VERSION : 1.1
// The function calculates a contour offset of a path (tool length and radius) / The function calculates a contour offset of a path (tool length and radius offset)
   VAR_INPUT
      toolLength : LReal;   // Tool length
      toolRadius : LReal;   // Tool radius
      pathPlane : Int;   // Path plane: XZ= 0, YZ=1, XY= 2
      compensationDirection : Int;   // Tool radius compensation direction: left=1, right = 0
   END_VAR
   VAR_IN_OUT
      pathDataIn : "LKinCtrl_typeCOffPathDataIn";   // Path data in
      pathDataOut : "LKinCtrl_typeCOffPathDataOut";   // Path dat out
   END_VAR
   VAR_TEMP
      internalNumber : DInt;   // Internal error position
      boCmdInPathPlane : Bool;   // Command in path plane
      pathDataDelete : "LKinCtrl_typeCOffPathDataOut";   // Delete data structure
      tempCurrentPoint : "LKinCtrl_typeCOff3DPoint";   // End point 1st command - current command
      tempCurrentPointPathPlane : "LKinCtrl_typeCOff3DPoint";   // End point 1st command - current command - path plane
      tempCurrentPointRadComp : "LKinCtrl_typeCOff3DPoint";   // End point 1st command - current command - radius compensated
      tempNextCmdIn : "LKinCtrl_typeCOffCmdInInternal";   // Next command input
      tempNextButOneCmdIn : "LKinCtrl_typeCOffCmdInInternal";   // Next but one command input
      tempNextCmdOut : "LKinCtrl_typeCOffCmdOutInternal";   // Next command output
      tempIntermediateCmdOut : "LKinCtrl_typeCOffCmdOutInternal";   // Intermediate command output
      tempNextButOneCmdOut : "LKinCtrl_typeCOffCmdOutInternal";   // Next but one command output
      tempToolRadiusComp : Bool;   // TRUE: tool radius compensation used
      tempToolLengthComp : Bool;   // TRUE: tool length compensation used
      tempRetValue : Word;   // Return value
      tempMuA : LReal;
      tempMuB : LReal;
      tempCornerType : Int;
      tempPa : "LKinCtrl_typeCOff3DPoint";
      tempPb : "LKinCtrl_typeCOff3DPoint";
      tempDistance1 : LReal;
      tempDistance2 : LReal;
      tempAngle : LReal;
      tempMod : DInt;
      tempPathChoice : DInt;
      tempNextCmdEndPointLevelled : "LKinCtrl_typeCOff3DPoint";
      tempNextCmdIntermediatePointLevelled : "LKinCtrl_typeCOff3DPoint";
      tempNextButOneStartPointOrthShiftedLevelled : "LKinCtrl_typeCOff3DPoint";
      tempNextButOneCmdStartPointOrthTangShiftedLevelled : "LKinCtrl_typeCOff3DPoint";
      tempNextCmdStartPointOrhtShiftLevelled : "LKinCtrl_typeCOff3DPoint";
      tempDirectionUncompensatedVec : "LKinCtrl_typeCOff3DPoint";
      tempDirectionCompensatedVec : "LKinCtrl_typeCOff3DPoint";
      tempDirectionUncompensatedUnitVec : "LKinCtrl_typeCOff3DPoint";
      tempDirectionCompensatedUnitVec : "LKinCtrl_typeCOff3DPoint";
      tempLengthCompensatedPointDifferenceVec : LReal;
   END_VAR
   // Ret_Val : Retrun data
   VAR CONSTANT
      COFF_TRANSITION_TOLERANCE : LReal := 0.2;   // Tolerance for additional circle - outer corner
      ERR_COFF_INVALID_TOOL_LENGTH : Word := 16#8301;   // Error - invalid tool length
      ERR_COFF_INVALID_TOOL_RADIUS : Word := 16#8302;   // Error - invalid tool radius
      ERR_COFF_INVALID_PATH_PLANE : Word := 16#8303;   // Error - invalid path plane
      ERR_COFF_INVALID_COMPENSATION_DIRECTION : Word := 16#8304;   // Error - invalid compensation direction
      ERR_COFF_FUNCTION_NOT_SUPPORTED : Word := 16#8305;   // Error - functionality not supported
      ERR_COFF_INVALID_COMMAND_TYPE : Word := 16#8306;   // Error - invalid command type
      ERR_COFF_INVALID_CIRCLE_MODE : Word := 16#8307;   // Error - invalid circle mode
      ERR_COFF_INVALID_PATH_PLANE_OF_CIRCULAR_CMD : Word := 16#8308;   // Error - invalid path plane of a circular command
      ERR_COFF_INVALID_PATH_CHOICE_OF_CIRCULAR_CMD : Word := 16#8309;   // Error - invalid path choice of circular command
      ERR_COFF_INTERNAL : Word := 16#830F;   // Error - internal
      ERR_COFF_VECTOR_LENGTH_ZERO : Word := 16#8310;   // Error - vector length is zero
      ERR_COFF_INVALID_ACOS_ARGUMENT : Word := 16#8311;   // Error - invalid ACOS argument
      ERR_COFF_LINES_DO_NOT_INTERSECT : Word := 16#8312;   // Error - no solution, lines don't intersect
      ERR_COFF_ZERO_VECTOR : Word := 16#8313;   // Error - zero vector
      ERR_COFF_CMD_LENGTH_ZERO : Word := 16#8314;   // Error - cmd with length zero not permitted
      ERR_COFF_LINE_CIRCLE_DO_NOT_INTERSECT : Word := 16#8315;   // Error - no solution - line and circle don't intersect
      ERR_COFF_CIRCLES_DO_NOT_INTERSECT : Word := 16#8318;   // Error - no solution - circles don't intersect
      ERR_COFF_ONE_CIRC_CONTAINED_IN_THE_OTHER : Word := 16#8319;   // Error - one circle is contained in the other
      ERR_COFF_NO_SOLUTION_FOR_GIVEN_LINEAR_CMD : Word := 16#8320;   // Error - no valid solution with given linear command
      ERR_COFF_NO_SOLUTION_FOR_GIVEN_CIRCULAR_CMD : Word := 16#8321;   // Error - no valid solution with given circular command
      ERR_COFF_LINEAR_CMD_AND_TOOL_RADIUS_LEAD_TO_REVERSAL : Word := 16#8322;   // Error - linear command in combination with tool radius leads to reversal movement / Error - no valid solution with given circular command
      ERR_COFF_CIRCLE_CENTERS_EQUAL : Word := 16#8350;   // Error - circle centers are equal infinite intersections (only internal)
      COFF_REGION_TYPE_NONE : Int := 0;   // Region type: none
      COFF_REGION_TYPE_PLAUSIBILITY : Int := 1;   // Region type: plausibitlity general
      COFF_REGION_TYPE_PLAUSIBILITY_NEXT_CMD : Int := 2;   // Region type: plausibility next command
      COFF_REGION_TYPE_PLAUSIBILITY_NEXT_BUT_ONE_CMD : Int := 3;   // Region type: plausibility next but one command
      COFF_REGION_TYPE_PRE_CALC : Int := 4;   // Region type: precalculation
      COFF_REGION_TYPE_RAD_COMP_NEXT_CMD_LIN : Int := 5;   // Region type: radius compensation next command linear
      COFF_REGION_TYPE_RAD_COMP_LIN_LIN : Int := 6;   // Region type: radius compensation next command linear, next but one command linear
      COFF_REGION_TYPE_RAD_COMP_LIN_CIRC : Int := 7;   // Region type: radius compensation next command linear, next but one command circular
      COFF_REGION_TYPE_RAD_COMP_LIN_NONE : Int := 8;   // Region type: radius compensation next command linear, next but one command none
      COFF_REGION_TYPE_RAD_COMP_LIN_GEN : Int := 9;   // Region type: radius compensation next command linear - general
      COFF_REGION_TYPE_RAD_COMP_NEXT_CMD_CIRC : Int := 10;   // Region type: radius compensation next command circular
      COFF_REGION_TYPE_RAD_COMP_CIRC_LIN : Int := 11;   // Region type: radius compensation next command circular next but one command linear
      COFF_REGION_TYPE_RAD_COMP_CIRC_CIRC : Int := 12;   // Region type: radius compensation next command circular, next but one command circular
      COFF_REGION_TYPE_RAD_COMP_CIRC_NONE : Int := 13;   // Region type: radius compensation next command circular, next but one command none
      COFF_REGION_TYPE_RAD_COMP_CIRC_GEN : Int := 14;   // Region type: radius compensation next command circular - general
      COFF_REGION_TYPE_LEN_COMP_NEXT : Int := 15;   // Region type: tool length compensation next command
      COFF_REGION_TYPE_LEN_COMP_INTER_CMD : Int := 16;   // Region type: tool length compensation intermediate command
      COFF_REGION_TYPE_LEN_COMP_NEXT_BUT_ONE_CMD : Int := 17;   // Region type: tool length compensation next but one command
      COFF_REGION_TYPE_OUTPUT_DATA : Int := 18;   // Region type: ouptut data
      COFF_TOLERANCE : LReal := 0.001;   // Tolerance
      COFF_CIRC_REVERSAL_TOLERANCE_ANGLE : LReal := 90.0;   // Reversal tolerance check for circle
   END_VAR
BEGIN
   //==========================================================================================
   // SIEMENS AG
   // (c)Copyright 2019 All Rights Reserved
   //------------------------------------------------------------------------------------------
   // Library: LKinCtrl
   // Tested with: S7-1515T-3 PN/DP
   // Engineering: TIA Portal V15
   // Restrictions: ---
   // Requirements: S7-1500T FW 2.5
   // Functionality: LKinCtrl_OffsetContour
   // The function calculates a contour offset of a path (tool length and radius) 
   // Support: tech.team.motioncontrol@siemens.com
   // Note: Parameter comments are only available in language 'English (United States)'
   //------------------------------------------------------------------------------------------
   // Change log table:
   // Version    Date          Expert in charge    Changes applied
   // 00.09.00   2019-02-06    AW                  // Beta version
   // 01.00.00   2019-03-08    AW                  // First release version
   // 01.01.00   2020-08-14    AW                  // Bug fix - intersection point of 1st and 2nd circle (equal circle centers)
   //                                              //         - LKinCtrl_CalcLineCircleIntersectionPoint
   //                                              //         - LKinCtrl_CalcCircleCircleIntersectionPoint
   //                                              // length compensation (circle with radius and endpoint)
   // 01.01.01  2020-08-25     AW                  // Additional tolerance intersection of two circles (possible tiny floating point
   //                                                 deviations in case of one intersection point) - LKinCtrl_CalcCircleCircleIntersectionPoint
   // 01.01.02  2020-10-13     AW                  // fix - check innter outer corner - not done for linear commands in same direction anymore
   //                                              // additional check for next command LINEAR and next but one command NONE
   //                                              // avoid reversal movement for small linear path length in combination with big compensation radius
   // 01.01.03  2020-11-09     AW                  // bugfix addtional check - N E X T   B U T   O N E   C M D  -  N O N E                                          
   //===========================================================================================

   // Plausibility checks of parameter
   REGION PLAUSIBILITY_CHECK
     // Check tool length
     IF (#toolLength < 0.0)
     THEN
       #LKinCtrl_OffsetContour.returnValue := #ERR_COFF_INVALID_TOOL_LENGTH; // Invalid tool length
       #LKinCtrl_OffsetContour."region" := #COFF_REGION_TYPE_PLAUSIBILITY;
       #LKinCtrl_OffsetContour.internalNumber := 101;
       RETURN;

     // Check tool radius  
     ELSIF (#toolRadius < 0.0)
     THEN
       #LKinCtrl_OffsetContour.returnValue := #ERR_COFF_INVALID_TOOL_RADIUS; // Invalid tool radius
       #LKinCtrl_OffsetContour."region" := #COFF_REGION_TYPE_PLAUSIBILITY;
       #LKinCtrl_OffsetContour.internalNumber := 102;
       RETURN;
     END_IF;

     // Check circular path plane in combination with global path plane - next command
     IF ((((#pathDataIn.nextCommand.cmdType = "LKINCTRL_MC_MOVECIRCULARABS") OR
       (#pathDataIn.nextCommand.cmdType = "LKINCTRL_MC_MOVECIRCULARREL")) AND
       ((#pathDataIn.nextCommand.cmdParameters.circleParameters.circMode = "CM_CENTER") OR
       (#pathDataIn.nextCommand.cmdParameters.circleParameters.circMode = "CM_RADIUS")) AND
       (#pathPlane <> #pathDataIn.nextCommand.cmdParameters.circleParameters.circlePlane)))
     THEN
       #LKinCtrl_OffsetContour.returnValue := #ERR_COFF_INVALID_PATH_PLANE_OF_CIRCULAR_CMD; // Invalid path plane of a circular command
       #LKinCtrl_OffsetContour."region" := #COFF_REGION_TYPE_PLAUSIBILITY_NEXT_CMD;
       #LKinCtrl_OffsetContour.internalNumber := 103;
       RETURN;
     END_IF;

     // Check circular path plane in combination with global path plane - next but one command
     IF((((#pathDataIn.nextButOneCommand.cmdType = "LKINCTRL_MC_MOVECIRCULARABS") OR
       (#pathDataIn.nextButOneCommand.cmdType = "LKINCTRL_MC_MOVECIRCULARREL")) AND
       ((#pathDataIn.nextButOneCommand.cmdParameters.circleParameters.circMode = "CM_CENTER") OR
       (#pathDataIn.nextButOneCommand.cmdParameters.circleParameters.circMode = "CM_RADIUS")) AND
       (#pathPlane <> #pathDataIn.nextButOneCommand.cmdParameters.circleParameters.circlePlane)))
     THEN
       #LKinCtrl_OffsetContour.returnValue := #ERR_COFF_INVALID_PATH_PLANE_OF_CIRCULAR_CMD; // Invalid path plane of a circular command
       #LKinCtrl_OffsetContour."region" := #COFF_REGION_TYPE_PLAUSIBILITY_NEXT_BUT_ONE_CMD;
       #LKinCtrl_OffsetContour.internalNumber := 104;
       RETURN;
     END_IF;

     // Tool radius compensation?
     #tempToolRadiusComp := FALSE;
     IF (#toolRadius > 0.0)
     THEN
       // Check path plane
       IF ((#pathPlane >= "CP_XZ") AND (#pathPlane <= "CP_XY"))
       THEN
         IF ((#compensationDirection >= "LKINCTRL_COMP_LEFT") AND (#compensationDirection <= "LKINCTRL_COMP_RIGHT"))
         THEN
           #tempToolRadiusComp := TRUE;
         ELSE
           #LKinCtrl_OffsetContour.returnValue := #ERR_COFF_INVALID_COMPENSATION_DIRECTION; // Invalid compensation direction
           #LKinCtrl_OffsetContour."region" := #COFF_REGION_TYPE_PLAUSIBILITY;
           #LKinCtrl_OffsetContour.internalNumber := 105;
           RETURN;
         END_IF;
       ELSE
         #LKinCtrl_OffsetContour.returnValue := #ERR_COFF_INVALID_PATH_PLANE; // Invalid path plane
         #LKinCtrl_OffsetContour."region" := #COFF_REGION_TYPE_PLAUSIBILITY;
         #LKinCtrl_OffsetContour.internalNumber := 106;
         RETURN;
       END_IF;
     END_IF;

     // Tool length compensation=
     IF (#toolLength > 0.0)
     THEN
       #tempToolLengthComp := TRUE;
     ELSE
       #tempToolLengthComp := FALSE;
     END_IF;
   END_REGION PLAUSIBILITY_CHECK


   REGION Delete data
     #pathDataOut := #pathDataDelete;
   END_REGION

   REGION General

     IF (#tempToolRadiusComp OR #tempToolLengthComp) THEN
       // Output data preliminary
       // Next command
       #pathDataOut.nextCommand := #pathDataIn.nextCommand;
       // Current position
       // --------------------------
       #tempCurrentPoint := "LKinCtrl_CartesianCoordTo3DPoint"(#pathDataIn.currentPos.positionAbsolute);
       #tempCurrentPointRadComp := "LKinCtrl_CartesianCoordTo3DPoint"(#pathDataIn.currentPos.positionAbsoluteRadComp);

       // Next command
       // --------------------------
       #tempNextCmdIn.cmdType := #pathDataIn.nextCommand.cmdType;
       // Write to output data - modifications done later
       #tempNextCmdOut.cmdType := #tempNextCmdIn.cmdType;

       #tempNextCmdIn.transitionParameter1 := #pathDataIn.nextCommand.cmdParameters.transitionParameters[1];
       #tempNextCmdIn.bufferMode := #pathDataIn.nextCommand.cmdParameters.bufferMode;

       IF ((#tempNextCmdIn.cmdType = "LKINCTRL_MC_MOVELINEARABS") OR
         (#tempNextCmdIn.cmdType = "LKINCTRL_MC_MOVELINEARREL"))
       THEN
         IF (#tempNextCmdIn.cmdType = "LKINCTRL_MC_MOVELINEARABS") THEN
           // Absolute coordinates
           // End point is defined

           #tempNextCmdIn.endPoint := "LKinCtrl_CartesianCoordTo3DPoint"(cartesianCoord := #pathDataIn.nextCommand.cmdCoordinates.cartesianPosition);

         ELSIF (#tempNextCmdIn.cmdType = "LKINCTRL_MC_MOVELINEARREL") THEN
           // Relative coordinates -> calculate absolute coordinate
           #tempNextCmdIn.endPoint := "LKinCtrl_VecAdd"(vIn1 := #tempCurrentPoint,
                                                        vIn2 := "LKinCtrl_CartesianCoordTo3DPoint"(#pathDataIn.nextCommand.cmdCoordinates.cartesianPosition));

           // Set command type to absolute
           #tempNextCmdOut.cmdType := "LKINCTRL_MC_MOVELINEARABS";
         END_IF;

         // Check if cmd length is unequal zero
         IF ("LKinCtrl_VecAbs"("LKinCtrl_VecSub"(vIn1 := #tempCurrentPoint, vIn2 := #tempNextCmdIn.endPoint)) < #COFF_TOLERANCE) THEN

           // Not allowed - function has no memory and therefore can't treat a command length of zero correctly
           #LKinCtrl_OffsetContour.returnValue := #ERR_COFF_CMD_LENGTH_ZERO;
           #LKinCtrl_OffsetContour."region" := #COFF_REGION_TYPE_PLAUSIBILITY_NEXT_CMD;
           #LKinCtrl_OffsetContour.internalNumber := 201;
           RETURN;
         END_IF;

         // Check if next linear command has at least one component in path plane direction
         #tempRetValue := "LKinCtrl_CalcVecDistancePathPlane"(vectorInA := #tempCurrentPoint,
                                                              vectorInB := #tempNextCmdIn.endPoint,
                                                              pathPlane := #pathPlane,
                                                              distancePathPlane => #tempDistance1);

         IF (#tempRetValue <> 0) THEN
           #LKinCtrl_OffsetContour.returnValue := #tempRetValue;
           #LKinCtrl_OffsetContour."region" := #COFF_REGION_TYPE_PLAUSIBILITY_NEXT_CMD;
           #LKinCtrl_OffsetContour.subBlockNumber := 35055;
           #LKinCtrl_OffsetContour.internalNumber := 202;
           RETURN;
         END_IF;

         // Check if movement is in respective path plane
         IF (#tempDistance1 > 0.0) THEN
           // Change current position?
           // --------------------------
           #boCmdInPathPlane := true;
         ELSE
           #boCmdInPathPlane := false;
         END_IF;

       ELSIF ((#tempNextCmdIn.cmdType = "LKINCTRL_MC_MOVECIRCULARABS") OR
         (#tempNextCmdIn.cmdType = "LKINCTRL_MC_MOVECIRCULARREL"))
       THEN

         #tempNextCmdIn.circleMode := #pathDataIn.nextCommand.cmdParameters.circleParameters.circMode;
         #tempNextCmdIn.pathChoice := #pathDataIn.nextCommand.cmdParameters.circleParameters.pathChoice;

         // Check for invalid path choice
         IF ((#tempNextCmdIn.pathChoice < "PC_POSITIVE") OR
           (#tempNextCmdIn.pathChoice > "PC_NEGATIVE"))
         THEN
           #LKinCtrl_OffsetContour.returnValue := #ERR_COFF_INVALID_PATH_CHOICE_OF_CIRCULAR_CMD; // Invalid path plane of a circular command
           #LKinCtrl_OffsetContour."region" := #COFF_REGION_TYPE_PLAUSIBILITY_NEXT_CMD;
           #LKinCtrl_OffsetContour.internalNumber := 203;
           RETURN;
         END_IF;

         #tempNextCmdIn.circlePlane := #pathDataIn.nextCommand.cmdParameters.circleParameters.circlePlane;

         IF ((#tempNextCmdIn.circleMode = "CM_BORDER") OR
           (#tempNextCmdIn.circleMode = "CM_RADIUS"))
         THEN
           // End point is defined
           IF (#tempNextCmdIn.cmdType = "LKINCTRL_MC_MOVECIRCULARABS") THEN
             // Absolute coordinates
             #tempNextCmdIn.endPoint := "LKinCtrl_CartesianCoordTo3DPoint"(cartesianCoord := #pathDataIn.nextCommand.cmdCoordinates.cartesianPosition);
           ELSE
             // Relative coordinates -> calculate absolute coordinate
             #tempNextCmdIn.endPoint := "LKinCtrl_VecAdd"(vIn1 := #tempCurrentPoint,
                                                          vIn2 := "LKinCtrl_CartesianCoordTo3DPoint"(#pathDataIn.nextCommand.cmdCoordinates.cartesianPosition));
           END_IF;

           IF (#tempNextCmdIn.circleMode = "CM_BORDER") THEN
             IF (#tempNextCmdIn.cmdType = "LKINCTRL_MC_MOVECIRCULARABS") THEN
               // Absolute coordinates
               #tempNextCmdIn.circleIntermediatePoint.x := #pathDataIn.nextCommand.cmdParameters.circleParameters.auxPoint[1];
               #tempNextCmdIn.circleIntermediatePoint.y := #pathDataIn.nextCommand.cmdParameters.circleParameters.auxPoint[2];
               #tempNextCmdIn.circleIntermediatePoint.z := #pathDataIn.nextCommand.cmdParameters.circleParameters.auxPoint[3];
             ELSE
               // Relative coordinates -> calculate absolute coordinate
               #tempNextCmdIn.circleIntermediatePoint.x := #tempCurrentPoint.x + #pathDataIn.nextCommand.cmdParameters.circleParameters.auxPoint[1];
               #tempNextCmdIn.circleIntermediatePoint.y := #tempCurrentPoint.y + #pathDataIn.nextCommand.cmdParameters.circleParameters.auxPoint[2];
               #tempNextCmdIn.circleIntermediatePoint.z := #tempCurrentPoint.z + #pathDataIn.nextCommand.cmdParameters.circleParameters.auxPoint[3];
             END_IF;
           END_IF;

           IF (#tempNextCmdIn.circleMode = "CM_RADIUS") THEN
             #tempNextCmdIn.circleRadius := #pathDataIn.nextCommand.cmdParameters.circleParameters.radius;

             // "Third" coordinate is ignored by system - also ignore here!
             // Use start coordinate of circle instead
             IF (#pathPlane = "CP_XZ") THEN
               #tempNextCmdIn.endPoint.y := #tempCurrentPoint.y;
             ELSIF (#pathPlane = "CP_YZ") THEN
               #tempNextCmdIn.endPoint.x := #tempCurrentPoint.x;
             ELSIF (#pathPlane = "CP_XY") THEN
               #tempNextCmdIn.endPoint.z := #tempCurrentPoint.z;
             END_IF;
           END_IF;

         ELSIF (#tempNextCmdIn.circleMode = "CM_CENTER") THEN
           #tempNextCmdIn.circleAngle := #pathDataIn.nextCommand.cmdParameters.circleParameters.arc;

           IF (#tempNextCmdIn.cmdType = "LKINCTRL_MC_MOVECIRCULARABS") THEN
             // Absolute coordinates
             #tempNextCmdIn.circleCenterPoint.x := #pathDataIn.nextCommand.cmdParameters.circleParameters.auxPoint[1];
             #tempNextCmdIn.circleCenterPoint.y := #pathDataIn.nextCommand.cmdParameters.circleParameters.auxPoint[2];
             #tempNextCmdIn.circleCenterPoint.z := #pathDataIn.nextCommand.cmdParameters.circleParameters.auxPoint[3];
           ELSE
             // Relative coordinates -> calculate absolute coordinate
             #tempNextCmdIn.circleCenterPoint.x := #tempCurrentPoint.x + #pathDataIn.nextCommand.cmdParameters.circleParameters.auxPoint[1];
             #tempNextCmdIn.circleCenterPoint.y := #tempCurrentPoint.y + #pathDataIn.nextCommand.cmdParameters.circleParameters.auxPoint[2];
             #tempNextCmdIn.circleCenterPoint.z := #tempCurrentPoint.z + #pathDataIn.nextCommand.cmdParameters.circleParameters.auxPoint[3];
           END_IF;
           IF (#tempNextCmdIn.circleMode = "CM_CENTER") THEN
             // "Third" coordinate is ignored by system - also ignore here!
             // Use start coordinate of circle instead
             IF (#pathPlane = "CP_XZ") THEN
               #tempNextCmdIn.circleCenterPoint.y := #tempCurrentPoint.y;
             ELSIF (#pathPlane = "CP_YZ") THEN
               #tempNextCmdIn.circleCenterPoint.x := #tempCurrentPoint.x;
             ELSIF (#pathPlane = "CP_XY") THEN
               #tempNextCmdIn.circleCenterPoint.z := #tempCurrentPoint.z;
             END_IF;

             // Calculte correct circle end point - parameter not mandatory (and therefore probably not correct)
             #tempRetValue := "LKinCtrl_CalcCircEndPointWithGivenCenterAndAngle"(circleStartPoint := #tempCurrentPoint,
                                                                                 circleCenterPoint := #tempNextCmdIn.circleCenterPoint,
                                                                                 pathPlane := #pathPlane,
                                                                                 pathChoice := #tempNextCmdIn.pathChoice,
                                                                                 angle := #tempNextCmdIn.circleAngle,
                                                                                 endPoint => #tempNextCmdIn.endPoint); // absolute coordinate

             IF (#tempRetValue <> 0) THEN
               #LKinCtrl_OffsetContour.returnValue := #tempRetValue;
               #LKinCtrl_OffsetContour."region" := #COFF_REGION_TYPE_PRE_CALC;
               #LKinCtrl_OffsetContour.subBlockNumber := 35053;
               #LKinCtrl_OffsetContour.internalNumber := 204;
               RETURN;
             END_IF;
           END_IF;

         ELSE
           #LKinCtrl_OffsetContour.returnValue := #ERR_COFF_INVALID_CIRCLE_MODE; // Invalid circle mode
           #LKinCtrl_OffsetContour."region" := #COFF_REGION_TYPE_PLAUSIBILITY_NEXT_CMD;
           RETURN;
         END_IF;

         // Set command type to absolute
         #tempNextCmdOut.cmdType := "LKINCTRL_MC_MOVECIRCULARABS";
       ELSE
         #LKinCtrl_OffsetContour.returnValue := #ERR_COFF_INVALID_COMMAND_TYPE; // Invalid command type
         #LKinCtrl_OffsetContour."region" := #COFF_REGION_TYPE_PLAUSIBILITY_NEXT_CMD;
         #LKinCtrl_OffsetContour.internalNumber := 205;
         RETURN;
       END_IF;

       // Write to output data - modifications done later
       #tempNextCmdOut.circleMode := #tempNextCmdIn.circleMode;
       #tempNextCmdOut.endPoint := #tempNextCmdIn.endPoint;
       #tempNextCmdOut.circleIntermediatePoint := #tempNextCmdIn.circleIntermediatePoint;
       #tempNextCmdOut.circleCenterPoint := #tempNextCmdIn.circleCenterPoint;
       #tempNextCmdOut.transitionParameter1 := #tempNextCmdIn.transitionParameter1;
       #tempNextCmdOut.circleAngle := #tempNextCmdIn.circleAngle;

       // Next but one command - important!
       #tempNextButOneCmdIn.transitionParameter1 := #pathDataIn.nextButOneCommand.cmdParameters.transitionParameters[1];
       #tempNextButOneCmdOut.transitionParameter1 := #tempNextButOneCmdIn.transitionParameter1;
     END_IF;
   END_REGION

   // Tool radius compensation
   REGION TOOL_RADIUS_COMPENSATION
     // Copy important source variables into temporary variables

     IF (#tempToolRadiusComp) THEN

       REGION Copy data
         // ############# C O P Y   D A T A #############
         // #################################### 

         // Next but one command
         //#pathDataOut.nextButOneCommand.transitionParameter := #pathDataIn.nextButOneCommand.cmdParameters.transitionParameters;

         // Next but one command
         // --------------------------
         #tempNextButOneCmdIn.cmdType := #pathDataIn.nextButOneCommand.cmdType;
         // Write to output data - modifications done later
         #tempNextButOneCmdOut.cmdType := #tempNextButOneCmdIn.cmdType;


         #tempNextButOneCmdIn.bufferMode := #pathDataIn.nextButOneCommand.cmdParameters.bufferMode;

         // End point is defined
         IF (#tempNextButOneCmdIn.cmdType = "LKINCTRL_MC_MOVELINEARABS") THEN
           // Absolute coordinates
           #tempNextButOneCmdIn.endPoint := "LKinCtrl_CartesianCoordTo3DPoint"(#pathDataIn.nextButOneCommand.cmdCoordinates.cartesianPosition);

         ELSIF (#tempNextButOneCmdIn.cmdType = "LKINCTRL_MC_MOVELINEARREL") THEN
           // Relative coordinates -> calculate absolute coordinate
           #tempNextButOneCmdIn.endPoint := "LKinCtrl_VecAdd"(vIn1 := #tempNextCmdIn.endPoint,
                                                              vIn2 := "LKinCtrl_CartesianCoordTo3DPoint"(#pathDataIn.nextButOneCommand.cmdCoordinates.cartesianPosition));

           // Set command type to absolute
           #tempNextButOneCmdOut.cmdType := "LKINCTRL_MC_MOVELINEARABS";

         ELSIF ((#tempNextButOneCmdIn.cmdType = "LKINCTRL_MC_MOVECIRCULARABS") OR
           (#tempNextButOneCmdIn.cmdType = "LKINCTRL_MC_MOVECIRCULARREL"))
         THEN
           #tempNextButOneCmdIn.circleMode := #pathDataIn.nextButOneCommand.cmdParameters.circleParameters.circMode;
           #tempNextButOneCmdIn.pathChoice := #pathDataIn.nextButOneCommand.cmdParameters.circleParameters.pathChoice;

           // Check for invalid path choice
           IF ((#tempNextButOneCmdIn.pathChoice < "PC_POSITIVE") OR
             (#tempNextButOneCmdIn.pathChoice > "PC_NEGATIVE"))
           THEN
             #LKinCtrl_OffsetContour.returnValue := #ERR_COFF_INVALID_PATH_CHOICE_OF_CIRCULAR_CMD; // Invalid path plane of a circular command
             #LKinCtrl_OffsetContour."region" := #COFF_REGION_TYPE_PLAUSIBILITY_NEXT_BUT_ONE_CMD;
             #LKinCtrl_OffsetContour.internalNumber := 210;
             RETURN;
           END_IF;

           #tempNextButOneCmdIn.circlePlane := #pathDataIn.nextButOneCommand.cmdParameters.circleParameters.circlePlane;

           IF ((#tempNextButOneCmdIn.circleMode = "CM_BORDER") OR
             (#tempNextButOneCmdIn.circleMode = "CM_RADIUS"))
           THEN

             // End point is defined
             IF (#tempNextButOneCmdIn.cmdType = "LKINCTRL_MC_MOVECIRCULARABS") THEN
               // Absolute coordinates
               #tempNextButOneCmdIn.endPoint := "LKinCtrl_CartesianCoordTo3DPoint"(#pathDataIn.nextButOneCommand.cmdCoordinates.cartesianPosition);
             ELSE
               // Relative coordinates -> calculate absolute coordinate 
               #tempNextButOneCmdIn.endPoint := "LKinCtrl_VecAdd"(vIn1 := #tempNextCmdIn.endPoint,
                                                                  vIn2 := "LKinCtrl_CartesianCoordTo3DPoint"(#pathDataIn.nextButOneCommand.cmdCoordinates.cartesianPosition));
             END_IF;

             IF (#tempNextButOneCmdIn.circleMode = "CM_BORDER") THEN
               IF (#tempNextButOneCmdIn.cmdType = "LKINCTRL_MC_MOVECIRCULARABS") THEN
                 // Absolute coordinates
                 #tempNextButOneCmdIn.circleIntermediatePoint.x := #pathDataIn.nextButOneCommand.cmdParameters.circleParameters.auxPoint[1];
                 #tempNextButOneCmdIn.circleIntermediatePoint.y := #pathDataIn.nextButOneCommand.cmdParameters.circleParameters.auxPoint[2];
                 #tempNextButOneCmdIn.circleIntermediatePoint.z := #pathDataIn.nextButOneCommand.cmdParameters.circleParameters.auxPoint[3];
               ELSE
                 // Relative coordinates -> calculate absolute coordinate
                 #tempNextButOneCmdIn.circleIntermediatePoint.x := #tempNextCmdIn.endPoint.x + #pathDataIn.nextButOneCommand.cmdParameters.circleParameters.auxPoint[1];
                 #tempNextButOneCmdIn.circleIntermediatePoint.y := #tempNextCmdIn.endPoint.y + #pathDataIn.nextButOneCommand.cmdParameters.circleParameters.auxPoint[2];
                 #tempNextButOneCmdIn.circleIntermediatePoint.z := #tempNextCmdIn.endPoint.z + #pathDataIn.nextButOneCommand.cmdParameters.circleParameters.auxPoint[3];
               END_IF;
             END_IF;

             IF (#tempNextButOneCmdIn.circleMode = "CM_RADIUS") THEN
               #tempNextButOneCmdIn.circleRadius := #pathDataIn.nextButOneCommand.cmdParameters.circleParameters.radius;

               // "Third" coordinate is ignored by system - also ignore here!
               // Use start coordinate of circle instead
               IF (#pathPlane = "CP_XZ") THEN
                 #tempNextButOneCmdIn.endPoint.y := #tempNextCmdIn.endPoint.y;
               ELSIF (#pathPlane = "CP_YZ") THEN
                 #tempNextButOneCmdIn.endPoint.x := #tempNextCmdIn.endPoint.x;
               ELSIF (#pathPlane = "CP_XY") THEN
                 #tempNextButOneCmdIn.endPoint.z := #tempNextCmdIn.endPoint.z;
               END_IF;

             END_IF;

           ELSIF (#tempNextButOneCmdIn.circleMode = "CM_CENTER") THEN
             #tempNextButOneCmdIn.circleAngle := #pathDataIn.nextButOneCommand.cmdParameters.circleParameters.arc;

             IF (#tempNextButOneCmdIn.cmdType = "LKINCTRL_MC_MOVECIRCULARABS") THEN
               // Absolute coordinates
               #tempNextButOneCmdIn.circleCenterPoint.x := #pathDataIn.nextButOneCommand.cmdParameters.circleParameters.auxPoint[1];
               #tempNextButOneCmdIn.circleCenterPoint.y := #pathDataIn.nextButOneCommand.cmdParameters.circleParameters.auxPoint[2];
               #tempNextButOneCmdIn.circleCenterPoint.z := #pathDataIn.nextButOneCommand.cmdParameters.circleParameters.auxPoint[3];
             ELSE
               // Relative coordinates -> calculate absolute coordinate
               #tempNextButOneCmdIn.circleCenterPoint.x := #tempNextCmdIn.endPoint.x + #pathDataIn.nextButOneCommand.cmdParameters.circleParameters.auxPoint[1];
               #tempNextButOneCmdIn.circleCenterPoint.y := #tempNextCmdIn.endPoint.y + #pathDataIn.nextButOneCommand.cmdParameters.circleParameters.auxPoint[2];
               #tempNextButOneCmdIn.circleCenterPoint.z := #tempNextCmdIn.endPoint.z + #pathDataIn.nextButOneCommand.cmdParameters.circleParameters.auxPoint[3];
             END_IF;

             // "Third" coordinate is ignored by system - also ignore here!
             // Use start coordinate of circle instead
             IF (#pathPlane = "CP_XZ") THEN
               #tempNextButOneCmdIn.circleCenterPoint.y := #tempNextCmdIn.endPoint.y;
             ELSIF (#pathPlane = "CP_YZ") THEN
               #tempNextButOneCmdIn.circleCenterPoint.x := #tempNextCmdIn.endPoint.x;
             ELSIF (#pathPlane = "CP_XY") THEN
               #tempNextButOneCmdIn.circleCenterPoint.z := #tempNextCmdIn.endPoint.z;
             END_IF;

           ELSE
             #LKinCtrl_OffsetContour.returnValue := #ERR_COFF_INVALID_CIRCLE_MODE; // Invalid circle mode
             #LKinCtrl_OffsetContour."region" := #COFF_REGION_TYPE_PLAUSIBILITY_NEXT_BUT_ONE_CMD;
             #LKinCtrl_OffsetContour.internalNumber := 211;
             RETURN;
           END_IF;

           // Set command type to absolute
           #tempNextButOneCmdOut.cmdType := "LKINCTRL_MC_MOVECIRCULARABS";

         ELSIF (#tempNextButOneCmdIn.cmdType = -1) THEN
           ;
         ELSE
           #LKinCtrl_OffsetContour.returnValue := #ERR_COFF_INVALID_COMMAND_TYPE; // Invalid command type
           #LKinCtrl_OffsetContour."region" := #COFF_REGION_TYPE_PLAUSIBILITY_NEXT_BUT_ONE_CMD;
           #LKinCtrl_OffsetContour.internalNumber := 212;
           RETURN;
         END_IF;

         // Write to output data - modifications done later
         #tempNextButOneCmdOut.circleMode := #tempNextButOneCmdIn.circleMode;
         #tempNextButOneCmdOut.endPoint := #tempNextButOneCmdIn.endPoint;
         #tempNextButOneCmdOut.circleIntermediatePoint := #tempNextButOneCmdIn.circleIntermediatePoint;
         #tempNextButOneCmdOut.circleCenterPoint := #tempNextButOneCmdIn.circleCenterPoint;


       END_REGION

       REGION Next command LINEAR

         // ############# N E X T   C M D  -  L I N E A R #############
         // ##############################################
         IF (#tempNextCmdOut.cmdType = "LKINCTRL_MC_MOVELINEARABS") THEN
           IF (#boCmdInPathPlane) THEN
             // ########## 1st linear command point 1 to point 2 ##########
             // Calculate tangential and orthogonal unit vector of direction
             #tempRetValue := "LKinCtrl_CalcLineTangOrthPathPlane"(pathPlane := #pathPlane,
                                                                   compDirection := #compensationDirection,
                                                                   vInFirst := #tempNextCmdIn.endPoint,
                                                                   vInSecond := #tempCurrentPoint,
                                                                   vUnitTangentialPathPlane => #tempNextCmdOut.tangentialUnitVecEnd,
                                                                   vUnitOrthogonalPathPlane => #tempNextCmdOut.orthogonalUnitVecEnd);

             IF (#tempRetValue <> 0) THEN
               #LKinCtrl_OffsetContour.returnValue := #tempRetValue;
               #LKinCtrl_OffsetContour."region" := #COFF_REGION_TYPE_RAD_COMP_NEXT_CMD_LIN;
               #LKinCtrl_OffsetContour.subBlockNumber := 35055;
               #LKinCtrl_OffsetContour.internalNumber := 301;
               RETURN;
             END_IF;

             // Scale othogonal vector with tool radius to get orthogonal shift
             #tempNextCmdOut.orthogonalShiftEnd := "LKinCtrl_VecScale"(vIn := #tempNextCmdOut.orthogonalUnitVecEnd,
                                                                       factor := #toolRadius);

             // Scale tangential vector with tool radius to get tangential shift
             #tempNextCmdOut.tangentiaShiftEnd := "LKinCtrl_VecScale"(vIn := #tempNextCmdOut.tangentialUnitVecEnd,
                                                                      factor := #toolRadius);

             // Calculate orthogonal shifted next target coordinate 
             #tempNextCmdOut.endPointOrthShifted := "LKinCtrl_VecAdd"(vIn1 := #tempNextCmdIn.endPoint,
                                                                      vIn2 := #tempNextCmdOut.orthogonalShiftEnd);

             // Calculate orthogonal and tangential shifted next target coordinate
             #tempNextCmdOut.endPointOrthTangShifted := "LKinCtrl_VecAdd"(vIn1 := #tempNextCmdOut.endPointOrthShifted,
                                                                          vIn2 := #tempNextCmdOut.tangentiaShiftEnd);

             #tempNextCmdOut.endPoint := #tempNextCmdOut.endPointOrthShifted;

             // ############# N E X T   B U T   O N E   C M D  -  L I N E A R #############
             IF (#tempNextButOneCmdOut.cmdType = "LKINCTRL_MC_MOVELINEARABS") THEN
               REGION Next but one command LINEAR
                 // 2nd linear command point 2 to point 3
                 // Calculate tangential and orthogonal unit vector of direction
                 #tempRetValue := "LKinCtrl_CalcLineTangOrthPathPlane"(pathPlane := #pathPlane,
                                                                       compDirection := #compensationDirection,
                                                                       vInFirst := #tempNextButOneCmdIn.endPoint,
                                                                       vInSecond := #tempNextCmdIn.endPoint,
                                                                       vUnitTangentialPathPlane => #tempNextButOneCmdOut.tangentialUnitVecStart,
                                                                       vUnitOrthogonalPathPlane => #tempNextButOneCmdOut.orthogonalUnitVecStart);

                 IF (#tempRetValue <> 0) THEN
                   #LKinCtrl_OffsetContour.returnValue := #tempRetValue;
                   #LKinCtrl_OffsetContour."region" := #COFF_REGION_TYPE_RAD_COMP_LIN_LIN;
                   #LKinCtrl_OffsetContour.subBlockNumber := 35055;
                   #LKinCtrl_OffsetContour.internalNumber := 302;
                   RETURN;
                 END_IF;

                 // Scale othogonal vector with tool radius to get orthogonal shift
                 #tempNextButOneCmdOut.orthogonalShiftStart := "LKinCtrl_VecScale"(vIn := #tempNextButOneCmdOut.orthogonalUnitVecStart,
                                                                                   factor := #toolRadius);

                 #tempNextButOneCmdOut.tangentiaShiftStart := "LKinCtrl_VecScale"(vIn := #tempNextButOneCmdOut.tangentialUnitVecStart,
                                                                                  factor := #toolRadius);

                 // Calculate orthogonal shifted next target coordinate 
                 #tempNextButOneCmdOut.startPointOrthShifted := "LKinCtrl_VecAdd"(vIn1 := #tempNextCmdIn.endPoint,
                                                                                  vIn2 := #tempNextButOneCmdOut.orthogonalShiftStart);

                 // Calculate orthogonal and tangential shifted next target coordinate
                 #tempNextButOneCmdOut.startPointOrthTangShifted := "LKinCtrl_VecAdd"(vIn1 := #tempNextButOneCmdOut.startPointOrthShifted,
                                                                                      vIn2 := #tempNextButOneCmdOut.tangentiaShiftStart);

                 // Check if 1st and 2nd linear command are located in exactly the same direction (tangential vector) - then orhtogonal shifted end point of next command is the solution!
                 // No intersection point, lines intersect completely!
                 #tempDistance1 := ("LKinCtrl_VecAbs"("LKinCtrl_VecSub"(vIn1 := #tempNextCmdOut.tangentialUnitVecEnd, vIn2 := #tempNextButOneCmdOut.tangentialUnitVecStart)));

                 // Check for zero vector
                 #tempDistance2 := ("LKinCtrl_VecAbs"(#tempNextButOneCmdOut.tangentialUnitVecStart));

                 IF ((#tempDistance1 > #COFF_TOLERANCE) AND (#tempDistance2 > 0.0)) THEN
                   // ########## Intersection point of 1st and 2nd linear command ##########
                   #tempRetValue := "LKinCtrl_CalcLineLineIntersectionPoint"(startPointFirstLine := #tempNextCmdOut.endPointOrthShifted,
                                                                             endPointFirstLine := #tempNextCmdOut.endPointOrthTangShifted,
                                                                             startPointSecondLine := #tempNextButOneCmdOut.startPointOrthShifted,
                                                                             endPointSecondLine := #tempNextButOneCmdOut.startPointOrthTangShifted,
                                                                             intersectionPointA => #tempPa,
                                                                             intersectionPointB => #tempPb,
                                                                             muA => #tempMuA,
                                                                             muB => #tempMuB);

                   IF (#tempRetValue <> 0) THEN
                     #LKinCtrl_OffsetContour.returnValue := #tempRetValue;
                     #LKinCtrl_OffsetContour."region" := #COFF_REGION_TYPE_RAD_COMP_LIN_LIN;
                     #LKinCtrl_OffsetContour.subBlockNumber := 35060;
                     #LKinCtrl_OffsetContour.internalNumber := 303;
                     RETURN;
                   END_IF;
                   #tempNextCmdOut.endPoint := #tempPa;
                 ELSE
                   #tempNextCmdOut.endPoint := #tempNextCmdOut.endPointOrthShifted;
                 END_IF;

                 // Check blending length
                 IF ((#tempNextButOneCmdIn.transitionParameter1 < 0.0) OR
                   // V01.01.02 AW 2020-10-13 - avoid inner / outer corner check if 1st and 2nd linear command are located in exactly the same direction
                   (#tempDistance1 < #COFF_TOLERANCE))
                 THEN
                   ; // Maximum blending length used - automatic algorithm, nothing to change here
                     // OR nothing to do - straight line
                 ELSE
                   // Distinguish between inner and outer corner
                   #tempRetValue := "LKinCtrl_CheckInnerOuterCorner"(vInFirst := #tempNextCmdOut.tangentialUnitVecEnd,
                                                                     vInSecond := #tempNextButOneCmdOut.tangentialUnitVecStart,
                                                                     pathPlane := #pathPlane,
                                                                     direction := #compensationDirection,
                                                                     cornerType => #tempCornerType);

                   IF (#tempRetValue <> 0) THEN
                     #LKinCtrl_OffsetContour.returnValue := #tempRetValue;
                     #LKinCtrl_OffsetContour."region" := #COFF_REGION_TYPE_RAD_COMP_LIN_LIN;
                     #LKinCtrl_OffsetContour.subBlockNumber := 35051;
                     #LKinCtrl_OffsetContour.internalNumber := 304;
                     RETURN;
                   END_IF;

                   IF (#tempCornerType = "LKINCTRL_OUTER_CORNER") THEN
                     IF (#tempNextButOneCmdIn.transitionParameter1 > #COFF_TRANSITION_TOLERANCE) THEN

                       // Output next but one coordinates - in case it's the last one
                       #tempNextButOneCmdOut.endPoint := "LKinCtrl_VecAdd"(vIn1 := #tempNextButOneCmdIn.endPoint,
                                                                           vIn2 := #tempNextButOneCmdOut.orthogonalShiftStart);


                       // Modify transition with blending distance - next but one command !
                       #tempNextButOneCmdOut.transitionParameter1 += #toolRadius;

                     ELSE
                       // Use shortened end point
                       #tempNextCmdOut.endPoint := #tempNextCmdOut.endPointOrthShifted;

                       // Additional command
                       // Intermediate command necessary (circle defined by intermediate position)
                       "LKinCtrl_CalcCircleIntermediatePos"(initialEndPoint := #tempNextCmdIn.endPoint,
                                                            newEndPoint := #tempPa,
                                                            toolRadius := #toolRadius,
                                                            circIntermediatePoint => #tempIntermediateCmdOut.circleIntermediatePoint);


                       #tempIntermediateCmdOut.cmdType := "LKINCTRL_MC_MOVECIRCULARABS";

                       #tempIntermediateCmdOut.endPoint := #tempNextButOneCmdOut.startPointOrthShifted;

                       // Definition via intermediate point and endpoint
                       #tempIntermediateCmdOut.circleMode := "CM_BORDER";

                     END_IF;
                   ELSE // Inner corner
                     ;
                   END_IF;
                 END_IF;
               END_REGION
               // #############  N E X T   B U T   O N E   C M D   -  C I R C U L A R #############
             ELSIF (#tempNextButOneCmdOut.cmdType = "LKINCTRL_MC_MOVECIRCULARABS") THEN
               REGION Next but one command CIRCULAR
                 // Use radius-compensated point (linear end point)
                 //#pathDataOut.nextCommand.cmdCoordinates.cartesianPosition := #tempNew2ndPoint;

                 // Distinguish between different circular modes
                 IF (#tempNextButOneCmdIn.circleMode = "CM_BORDER") THEN

                   // ------------ Via an intermediate point and the end point ("CircMode" = 0) ------------

                   // Caluclate center point of circle with given start point, end point and intermediate point
                   #tempRetValue := "LKinCtrl_CalcCircCenterByIntermediatePointAndEndPoint"(circleStartPoint := #tempNextCmdIn.endPoint,
                                                                                            circleEndPoint := #tempNextButOneCmdIn.endPoint,
                                                                                            circleIntermediatePoint := #tempNextButOneCmdIn.circleIntermediatePoint,
                                                                                            pathPlane := #pathPlane,
                                                                                            circleCenterPoint => #tempNextButOneCmdIn.circleCenterPoint);

                   IF (#tempRetValue <> 0) THEN
                     #LKinCtrl_OffsetContour.returnValue := #tempRetValue;
                     #LKinCtrl_OffsetContour."region" := #COFF_REGION_TYPE_RAD_COMP_LIN_CIRC;
                     #LKinCtrl_OffsetContour.subBlockNumber := 35057;
                     #LKinCtrl_OffsetContour.internalNumber := 330;
                     RETURN;
                   END_IF;

                   // Calculate path choice
                   #tempRetValue := "LKinCtrl_CalcCircPathChoiceByIntermediatePointAndEndPoint"(circleStartPoint := #tempNextCmdIn.endPoint,
                                                                                                circleEndPoint := #tempNextButOneCmdIn.endPoint,
                                                                                                circleintermediatePoint := #tempNextButOneCmdIn.circleIntermediatePoint,
                                                                                                pathPlane := #pathPlane,
                                                                                                pathChoice => #tempNextButOneCmdIn.pathChoice);


                   IF (#tempRetValue <> 0) THEN
                     #LKinCtrl_OffsetContour.returnValue := #tempRetValue;
                     #LKinCtrl_OffsetContour."region" := #COFF_REGION_TYPE_RAD_COMP_LIN_CIRC;
                     #LKinCtrl_OffsetContour.subBlockNumber := 35058;
                     #LKinCtrl_OffsetContour.internalNumber := 331;
                     RETURN;
                   END_IF;

                 ELSIF (#tempNextButOneCmdIn.circleMode = "CM_CENTER") THEN
                   // ------------ Via the circle center and the angle in a main plane ("CircMode" = 1) ------------
                   // "Third" coordinate is ignored by system - also ignore here!

                   // Calculte correct circle end point - parameter not mandatory (and therefore probably not correct)
                   #tempRetValue := "LKinCtrl_CalcCircEndPointWithGivenCenterAndAngle"(circleStartPoint := #tempNextCmdIn.endPoint,
                                                                                       circleCenterPoint := #tempNextButOneCmdIn.circleCenterPoint,
                                                                                       pathPlane := #pathPlane,
                                                                                       pathChoice := #tempNextButOneCmdIn.pathChoice,
                                                                                       angle := #tempNextButOneCmdIn.circleAngle,
                                                                                       endPoint => #tempNextButOneCmdIn.endPoint);




                   IF (#tempRetValue <> 0) THEN
                     #LKinCtrl_OffsetContour.returnValue := #tempRetValue;
                     #LKinCtrl_OffsetContour."region" := #COFF_REGION_TYPE_RAD_COMP_CIRC_CIRC;
                     #LKinCtrl_OffsetContour.subBlockNumber := 35053;
                     #LKinCtrl_OffsetContour.internalNumber := 332;
                     RETURN;
                   END_IF;

                 ELSIF (#tempNextButOneCmdIn.circleMode = "CM_RADIUS") THEN

                   // Calculate circle center point by given start / end point and radius and path choice
                   #tempRetValue := "LKinCtrl_CalcCircCenterByRadiusAndEndPoint"(circleStartPoint := #tempNextCmdIn.endPoint,
                                                                                 circleEndPoint := #tempNextButOneCmdIn.endPoint,
                                                                                 pathPlane := #pathPlane,
                                                                                 circleRadius := #tempNextButOneCmdIn.circleRadius,
                                                                                 pathChoice := #tempNextButOneCmdIn.pathChoice,
                                                                                 circCenterPoint => #tempNextButOneCmdIn.circleCenterPoint);

